   AddressMH[3].Ref_PLC_set_value_CP := 0;
   AddressMH[3].Ref_NozzelBypassControl := 0;
   AddressMH[3].Ref_NozzelBypassSetOut := 0;
   AddressMH[3].Ref_Reserve := 0;
   AddressMH[3].Ref_OK := FALSE;
   AddressMH[3].MH_Channel_01 := TRUE;
   AddressMH[3].MH_Channel_02 := FALSE;
   AddressMH[3].Spare_03 := FALSE;
   AddressMH[3].Spare_04 := FALSE;
   AddressMH[3].Spare_05 := FALSE;
   AddressMH[3].Spare_06 := FALSE;
   AddressMH[3].Spare_07 := FALSE;
   AddressMH[4].Ref_Digital_Input := 32;
   AddressMH[4].Ref_MH_ShotTime := 1550;
   AddressMH[4].Ref_MH_Opening_Time := 1554;
   AddressMH[4].Ref_MH_Closing_Time := 1556;
   AddressMH[4].Ref_MH_State := 1560;
   AddressMH[4].Ref_PLC_State := 0;
   AddressMH[4].Ref_CP_State := 0;
   AddressMH[4].Ref_Digital_Output := 32;
   AddressMH[4].Ref_ShotTimeSetValue := 1550;
   AddressMH[4].Ref_ServiceProduction := 1554;
   AddressMH[4].Ref_MixingheadControl := 1560;
   AddressMH[4].Ref_PLC_comand_SP := 0;
   AddressMH[4].Ref_PLC_comand_CP := 0;
   AddressMH[4].Ref_PLC_set_value_SP := 0;
   AddressMH[4].Ref_PLC_set_value_CP := 0;
   AddressMH[4].Ref_NozzelBypassControl := 0;
   AddressMH[4].Ref_NozzelBypassSetOut := 0;
   AddressMH[4].Ref_Reserve := 0;
   AddressMH[4].Ref_OK := FALSE;
   AddressMH[4].MH_Channel_01 := TRUE;
   AddressMH[4].MH_Channel_02 := FALSE;
   AddressMH[4].Spare_03 := FALSE;
   AddressMH[4].Spare_04 := FALSE;
   AddressMH[4].Spare_05 := FALSE;
   AddressMH[4].Spare_06 := FALSE;
   AddressMH[4].Spare_07 := FALSE;
   AddressMH[5].Ref_Digital_Input := 36;
   AddressMH[5].Ref_MH_ShotTime := 1636;
   AddressMH[5].Ref_MH_Opening_Time := 1640;
   AddressMH[5].Ref_MH_Closing_Time := 1642;
   AddressMH[5].Ref_MH_State := 1644;
   AddressMH[5].Ref_PLC_State := 0;
   AddressMH[5].Ref_CP_State := 0;
   AddressMH[5].Ref_Digital_Output := 36;
   AddressMH[5].Ref_ShotTimeSetValue := 1636;
   AddressMH[5].Ref_ServiceProduction := 1640;
   AddressMH[5].Ref_MixingheadControl := 1642;
   AddressMH[5].Ref_PLC_comand_SP := 0;
   AddressMH[5].Ref_PLC_comand_CP := 0;
   AddressMH[5].Ref_PLC_set_value_SP := 0;
   AddressMH[5].Ref_PLC_set_value_CP := 0;
   AddressMH[5].Ref_NozzelBypassControl := 0;
   AddressMH[5].Ref_NozzelBypassSetOut := 0;
   AddressMH[5].Ref_Reserve := 0;
   AddressMH[5].Ref_OK := FALSE;
   AddressMH[5].MH_Channel_01 := TRUE;
   AddressMH[5].MH_Channel_02 := FALSE;
   AddressMH[5].Spare_03 := FALSE;
   AddressMH[5].Spare_04 := FALSE;
   AddressMH[5].Spare_05 := FALSE;
   AddressMH[5].Spare_06 := FALSE;
   AddressMH[5].Spare_07 := FALSE;
   AddressMH[6].Ref_Digital_Input := 40;
   AddressMH[6].Ref_MH_ShotTime := 1686;
   AddressMH[6].Ref_MH_Opening_Time := 1690;
   AddressMH[6].Ref_MH_Closing_Time := 1692;
   AddressMH[6].Ref_MH_State := 1694;
   AddressMH[6].Ref_PLC_State := 0;
   AddressMH[6].Ref_CP_State := 0;
   AddressMH[6].Ref_Digital_Output := 40;
   AddressMH[6].Ref_ShotTimeSetValue := 1686;
   AddressMH[6].Ref_ServiceProduction := 1690;
   AddressMH[6].Ref_MixingheadControl := 1692;
   AddressMH[6].Ref_PLC_comand_SP := 0;
   AddressMH[6].Ref_PLC_comand_CP := 0;
   AddressMH[6].Ref_PLC_set_value_SP := 0;
   AddressMH[6].Ref_PLC_set_value_CP := 0;
   AddressMH[6].Ref_NozzelBypassControl := 0;
   AddressMH[6].Ref_NozzelBypassSetOut := 0;
   AddressMH[6].Ref_Reserve := 0;
   AddressMH[6].Ref_OK := FALSE;
   AddressMH[6].MH_Channel_01 := TRUE;
   AddressMH[6].MH_Channel_02 := FALSE;
   AddressMH[6].Spare_03 := FALSE;
   AddressMH[6].Spare_04 := FALSE;
   AddressMH[6].Spare_05 := FALSE;
   AddressMH[6].Spare_06 := FALSE;
   AddressMH[6].Spare_07 := FALSE;
   AddressMH[7].Ref_Digital_Input := 44;
   AddressMH[7].Ref_MH_ShotTime := 1736;
   AddressMH[7].Ref_MH_Opening_Time := 1740;
   AddressMH[7].Ref_MH_Closing_Time := 1742;
   AddressMH[7].Ref_MH_State := 1744;
   AddressMH[7].Ref_PLC_State := 0;
   AddressMH[7].Ref_CP_State := 0;
   AddressMH[7].Ref_Digital_Output := 44;
   AddressMH[7].Ref_ShotTimeSetValue := 1736;
   AddressMH[7].Ref_ServiceProduction := 1740;
   AddressMH[7].Ref_MixingheadControl := 1742;
   AddressMH[7].Ref_PLC_comand_SP := 0;
   AddressMH[7].Ref_PLC_comand_CP := 0;
   AddressMH[7].Ref_PLC_set_value_SP := 0;
   AddressMH[7].Ref_PLC_set_value_CP := 0;
   AddressMH[7].Ref_NozzelBypassControl := 0;
   AddressMH[7].Ref_NozzelBypassSetOut := 0;
   AddressMH[7].Ref_Reserve := 0;
   // 242 more start values not shown
END_DATA_BLOCK

DATA_BLOCK "DB1233_ProCanIO_Flow"   // DB1233
TITLE = Address allocation flow IO-ProCan
{ S7_Optimized_Access := 'FALSE' }
VERSION : 0.1
   VAR
      ReadWriteDeviceNo : Int := 1;
      CopyDeviceNO : Int := 0;
      Read : Bool := FALSE;
      Write : Bool := FALSE;
      Copy : Bool := FALSE;
      AddressFlow : Array[0..16] of "UDT1233_ProCanIO_Flow";
   END_VAR
BEGIN
   AddressFlow[1].Ref_Act_FlowValue := 2000;
   AddressFlow[2].Ref_Act_FlowValue := 2004;
   AddressFlow[3].Ref_Act_FlowValue := 800;
   AddressFlow[4].Ref_Act_FlowValue := 0;
   AddressFlow[5].Ref_Act_FlowValue := 0;
   AddressFlow[6].Ref_Act_FlowValue := 0;
   AddressFlow[7].Ref_Act_FlowValue := 0;
   AddressFlow[8].Ref_Act_FlowValue := 0;
   AddressFlow[9].Ref_Act_FlowValue := 0;
   AddressFlow[10].Ref_Act_FlowValue := 0;
   AddressFlow[11].Ref_Act_FlowValue := 0;
   AddressFlow[12].Ref_Act_FlowValue := 0;
   AddressFlow[1].Ref_Act_FlowState := 2032;
   AddressFlow[2].Ref_Act_FlowState := 2033;
   AddressFlow[3].Ref_Act_FlowState := 0;
   AddressFlow[4].Ref_Act_FlowState := 0;
   AddressFlow[5].Ref_Act_FlowState := 0;
   AddressFlow[6].Ref_Act_FlowState := 0;
   AddressFlow[7].Ref_Act_FlowState := 0;
   AddressFlow[8].Ref_Act_FlowState := 0;
   AddressFlow[9].Ref_Act_FlowState := 0;
   AddressFlow[10].Ref_Act_FlowState := 0;
   AddressFlow[11].Ref_Act_FlowState := 0;
   AddressFlow[12].Ref_Act_FlowState := 0;
   AddressFlow[1].Ref_Set_FlowRate := 2000;
   AddressFlow[2].Ref_Set_FlowRate := 2004;
   AddressFlow[3].Ref_Set_FlowRate := 0;
   AddressFlow[4].Ref_Set_FlowRate := 0;
   AddressFlow[5].Ref_Set_FlowRate := 0;
   AddressFlow[6].Ref_Set_FlowRate := 0;
   AddressFlow[7].Ref_Set_FlowRate := 0;
   AddressFlow[8].Ref_Set_FlowRate := 0;
   AddressFlow[9].Ref_Set_FlowRate := 0;
   AddressFlow[10].Ref_Set_FlowRate := 0;
   AddressFlow[11].Ref_Set_FlowRate := 0;
   AddressFlow[12].Ref_Set_FlowRate := 0;
   AddressFlow[1].Ref_Set_FlowRateQPB := 2016;
   AddressFlow[2].Ref_Set_FlowRateQPB := 2020;
   AddressFlow[3].Ref_Set_FlowRateQPB := 0;
   AddressFlow[4].Ref_Set_FlowRateQPB := 0;
   AddressFlow[5].Ref_Set_FlowRateQPB := 0;
   AddressFlow[6].Ref_Set_FlowRateQPB := 0;
   AddressFlow[7].Ref_Set_FlowRateQPB := 0;
   AddressFlow[8].Ref_Set_FlowRateQPB := 0;
   AddressFlow[9].Ref_Set_FlowRateQPB := 0;
   AddressFlow[10].Ref_Set_FlowRateQPB := 0;
   AddressFlow[11].Ref_Set_FlowRateQPB := 0;
   AddressFlow[12].Ref_Set_FlowRateQPB := 0;
   AddressFlow[1].Ref_Set_SWO_PressureQPB := 2032;
   AddressFlow[2].Ref_Set_SWO_PressureQPB := 2034;
   AddressFlow[3].Ref_Set_SWO_PressureQPB := 0;
   AddressFlow[4].Ref_Set_SWO_PressureQPB := 0;
   AddressFlow[5].Ref_Set_SWO_PressureQPB := 0;
   AddressFlow[6].Ref_Set_SWO_PressureQPB := 0;
   AddressFlow[7].Ref_Set_SWO_PressureQPB := 0;
   AddressFlow[8].Ref_Set_SWO_PressureQPB := 0;
   AddressFlow[9].Ref_Set_SWO_PressureQPB := 0;
   AddressFlow[10].Ref_Set_SWO_PressureQPB := 0;
   AddressFlow[11].Ref_Set_SWO_PressureQPB := 0;
   AddressFlow[12].Ref_Set_SWO_PressureQPB := 0;
   AddressFlow[1].Ref_Set_FlowIndexFlags := 2040;
   AddressFlow[2].Ref_Set_FlowIndexFlags := 2041;
   AddressFlow[3].Ref_Set_FlowIndexFlags := 0;
   AddressFlow[4].Ref_Set_FlowIndexFlags := 0;
   AddressFlow[5].Ref_Set_FlowIndexFlags := 0;
   AddressFlow[6].Ref_Set_FlowIndexFlags := 0;
   AddressFlow[7].Ref_Set_FlowIndexFlags := 0;
   AddressFlow[8].Ref_Set_FlowIndexFlags := 0;
   AddressFlow[9].Ref_Set_FlowIndexFlags := 0;
   AddressFlow[10].Ref_Set_FlowIndexFlags := 0;
   AddressFlow[11].Ref_Set_FlowIndexFlags := 0;
   AddressFlow[12].Ref_Set_FlowIndexFlags := 0;
   AddressFlow[1].Ref_PistonPosition := 0;
   AddressFlow[7].Ref_PistonPosition := 0;
   AddressFlow[1].Ref_OK := TRUE;
   AddressFlow[2].Ref_OK := TRUE;
   AddressFlow[3].Ref_OK := FALSE;
   AddressFlow[4].Ref_OK := FALSE;
   AddressFlow[5].Ref_OK := FALSE;
   AddressFlow[6].Ref_OK := FALSE;
   AddressFlow[7].Ref_OK := FALSE;
   AddressFlow[8].Ref_OK := FALSE;
   AddressFlow[9].Ref_OK := FALSE;
   AddressFlow[10].Ref_OK := FALSE;
   AddressFlow[11].Ref_OK := FALSE;
   AddressFlow[12].Ref_OK := FALSE;
   AddressFlow[3].Ref_Act_PressureQPB := 0;
   AddressFlow[3].Ref_TandemStatus := 0;
   AddressFlow[0].Ref_Act_FlowValue := 2000;
   AddressFlow[0].Ref_Act_FlowState := 2032;
   AddressFlow[0].Ref_Set_FlowRate := 2000;
   AddressFlow[0].Ref_Set_FlowRateQPB := 2016;
   AddressFlow[0].Ref_Act_PressureQPB := 0;
   AddressFlow[0].Ref_Set_SWO_PressureQPB := 2032;
   AddressFlow[0].Ref_Set_FlowIndexFlags := 2040;
   AddressFlow[0].Ref_TandemStatus := 0;
   AddressFlow[0].Ref_TandemComand := 0;
   AddressFlow[0].Ref_PistonPosition := 0;
   AddressFlow[0].Ref_OK := TRUE;
   AddressFlow[1].Ref_Act_PressureQPB := 0;
   AddressFlow[1].Ref_TandemStatus := 0;
   AddressFlow[1].Ref_TandemComand := 0;
   AddressFlow[2].Ref_Act_PressureQPB := 0;
   AddressFlow[2].Ref_TandemStatus := 0;
   AddressFlow[2].Ref_TandemComand := 0;
   AddressFlow[2].Ref_PistonPosition := 0;
   AddressFlow[3].Ref_TandemComand := 0;
   AddressFlow[3].Ref_PistonPosition := 0;
   AddressFlow[4].Ref_Act_PressureQPB := 0;
   AddressFlow[4].Ref_TandemStatus := 0;
   AddressFlow[4].Ref_TandemComand := 0;
   AddressFlow[4].Ref_PistonPosition := 0;
   AddressFlow[5].Ref_Act_PressureQPB := 0;
   AddressFlow[5].Ref_TandemStatus := 0;
   AddressFlow[5].Ref_TandemComand := 0;
   AddressFlow[5].Ref_PistonPosition := 0;
   AddressFlow[6].Ref_Act_PressureQPB := 0;
   AddressFlow[6].Ref_TandemStatus := 0;
   AddressFlow[6].Ref_TandemComand := 0;
   AddressFlow[6].Ref_PistonPosition := 0;
   AddressFlow[7].Ref_Act_PressureQPB := 0;
   AddressFlow[7].Ref_TandemStatus := 0;
   AddressFlow[7].Ref_TandemComand := 0;
   AddressFlow[8].Ref_Act_PressureQPB := 0;
   AddressFlow[8].Ref_TandemStatus := 0;
   AddressFlow[8].Ref_TandemComand := 0;
   AddressFlow[8].Ref_PistonPosition := 0;
   AddressFlow[9].Ref_Act_PressureQPB := 0;
   AddressFlow[9].Ref_TandemStatus := 0;
   AddressFlow[9].Ref_TandemComand := 0;
   AddressFlow[9].Ref_PistonPosition := 0;
   AddressFlow[10].Ref_Act_PressureQPB := 0;
   AddressFlow[10].Ref_TandemStatus := 0;
   AddressFlow[10].Ref_TandemComand := 0;
   AddressFlow[10].Ref_PistonPosition := 0;
   AddressFlow[11].Ref_Act_PressureQPB := 0;
   AddressFlow[11].Ref_TandemStatus := 0;
   AddressFlow[11].Ref_TandemComand := 0;
   AddressFlow[11].Ref_PistonPosition := 0;
   AddressFlow[12].Ref_Act_PressureQPB := 0;
   AddressFlow[12].Ref_TandemStatus := 0;
   AddressFlow[12].Ref_TandemComand := 0;
   AddressFlow[12].Ref_PistonPosition := 0;
   AddressFlow[13].Ref_Act_FlowValue := 0;
   AddressFlow[13].Ref_Act_FlowState := 0;
   AddressFlow[13].Ref_Set_FlowRate := 0;
   AddressFlow[13].Ref_Set_FlowRateQPB := 0;
   AddressFlow[13].Ref_Act_PressureQPB := 0;
   AddressFlow[13].Ref_Set_SWO_PressureQPB := 0;
   AddressFlow[13].Ref_Set_FlowIndexFlags := 0;
   AddressFlow[13].Ref_TandemStatus := 0;
   AddressFlow[13].Ref_TandemComand := 0;
   AddressFlow[13].Ref_PistonPosition := 0;
   AddressFlow[13].Ref_OK := FALSE;
   AddressFlow[14].Ref_Act_FlowValue := 0;
   AddressFlow[14].Ref_Act_FlowState := 0;
   AddressFlow[14].Ref_Set_FlowRate := 0;
   AddressFlow[14].Ref_Set_FlowRateQPB := 0;
   AddressFlow[14].Ref_Act_PressureQPB := 0;
   AddressFlow[14].Ref_Set_SWO_PressureQPB := 0;
   AddressFlow[14].Ref_Set_FlowIndexFlags := 0;
   AddressFlow[14].Ref_TandemStatus := 0;
   AddressFlow[14].Ref_TandemComand := 0;
   AddressFlow[14].Ref_PistonPosition := 0;
   AddressFlow[14].Ref_OK := FALSE;
   AddressFlow[15].Ref_Act_FlowValue := 0;
   AddressFlow[15].Ref_Act_FlowState := 0;
   AddressFlow[15].Ref_Set_FlowRate := 0;
   AddressFlow[15].Ref_Set_FlowRateQPB := 0;
   AddressFlow[15].Ref_Act_PressureQPB := 0;
   AddressFlow[15].Ref_Set_SWO_PressureQPB := 0;
   AddressFlow[15].Ref_Set_FlowIndexFlags := 0;
   AddressFlow[15].Ref_TandemStatus := 0;
   AddressFlow[15].Ref_TandemComand := 0;
   AddressFlow[15].Ref_PistonPosition := 0;
   AddressFlow[15].Ref_OK := FALSE;
   AddressFlow[16].Ref_Act_FlowValue := 0;
   AddressFlow[16].Ref_Act_FlowState := 0;
   AddressFlow[16].Ref_Set_FlowRate := 0;
   AddressFlow[16].Ref_Set_FlowRateQPB := 0;
   AddressFlow[16].Ref_Act_PressureQPB := 0;
   AddressFlow[16].Ref_Set_SWO_PressureQPB := 0;
   AddressFlow[16].Ref_Set_FlowIndexFlags := 0;
   AddressFlow[16].Ref_TandemStatus := 0;
   AddressFlow[16].Ref_TandemComand := 0;
   AddressFlow[16].Ref_PistonPosition := 0;
   AddressFlow[16].Ref_OK := FALSE;
END_DATA_BLOCK

DATA_BLOCK "DB1500_ShotDataToMC"   // DB1500
{ S7_Optimized_Access := 'FALSE' }
VERSION : 0.1
   VAR
      ShotData_MC : Array[0..4] of "ShotDataToMC";
   END_VAR
BEGIN
END_DATA_BLOCK

DATA_BLOCK "DB1900_IF_Robots"   // DB1900
{ S7_Optimized_Access := 'FALSE' }
VERSION : 0.1
   VAR
      ReadWriteDeviceNo : Int := 1;
      CopyDeviceNO : Int := 0;
      Read : Bool := FALSE;
      Write : Bool := FALSE;
      Copy : Bool := FALSE;
      Switch_Robots : Array[0..4] of Struct   // Switch Robots / State Robots
         SwitchHomePosON_OFF : Bool;
         SwitchMaintPosON_OFF : Bool;
         SwitchMaintPos_2ON_OFF : Bool;
         SwitchTestShotON_OFF : Bool;
         SwitchCleaningON_OFF : Bool;
         SwitchBrushON_OFF : Bool;
         SwitchSyncON_OFF : Bool;
         SwitchTeachenON_OFF : Bool;
         SwitchLearningON_OFF : Bool;
         SwitchAirCleaningON_OFF : Bool;
         SwitchAirCleaningManON_OFF : Bool;
         SwitchSpare_12 : Bool;
         SwitchSpare_13 : Bool;
         SwitchSpare_14 : Bool;
         SwitchSpare_15 : Bool;
         SwitchSpare_16 : Bool;
         StateHomePos : Byte;
         StateMaintPos : Byte;
         StateMaintPos_2 : Byte;
         StateTestShot : Byte;
         StateCleaning : Byte;
         StateBrush : Byte;
         StateSync : Byte;
         StateTeachen : Byte;
         StateLearning : Byte;
         StateAirCleaning : Byte;
         StateAirCleaningManual : Byte;
         State_12 : Byte;
         State_13 : Byte;
         State_14 : Byte;
         State_15 : Byte;
         State_16 : Byte;
      END_STRUCT;
      State_Robots : Array[0..4] of Struct   // State Robots for HMI
         Rob_in_Home : Bool;
         Rob_in_Automatic : Bool;
         Rob_in_Cycle : Bool;
         Fault_Exist : Bool;
         EmergencyStopReady : Bool;
         AutomatcStopReady : Bool;
         MixingheadAuto : Bool;
         MaschineAuto : Bool;
         CleaningMHRequested : Bool;
         CleaningMHOn : Bool;
         ReadyForStartCycle : Bool;
         TestShotRunning : Bool;
         AtPos1or2 : Bool;   // Die Schnittstellen an diesen Roboter sind an erster oder zweiter Stelle angemeldet
         Spare_1_5 : Bool;
         Spare_1_6 : Bool;
         Spare_1_7 : Bool;
         Rob_Prog_No : Byte;
         Rob_MC_No : Byte;
         StepNo : Byte;
         FaultNo : Byte;
         Spare_6 : Byte;
         Spare_7 : Byte;
         Spare_8 : Byte;
      END_STRUCT;
      Faults_Robots : Array[0..4] of "General_Faults";   // Faults Robots for HMI
      State_Kuka : Array[0..4] of "Kuka_KRC4_Status";   // State/Input/Ouput Kuka
      State_ABB : Array[0..4] of "ABB_IRC6_State";   // State/Input/Ouput ABB
      State_Fanuc : Array[0..4] of "Fanuc_Status";   // State/Input/Ouput Fanuc
   END_VAR
BEGIN
   Switch_Robots[0].SwitchHomePosON_OFF := FALSE;
   Switch_Robots[0].SwitchMaintPosON_OFF := FALSE;
   Switch_Robots[0].SwitchMaintPos_2ON_OFF := FALSE;
   Switch_Robots[0].SwitchTestShotON_OFF := FALSE;
   Switch_Robots[0].SwitchCleaningON_OFF := FALSE;
   Switch_Robots[0].SwitchBrushON_OFF := FALSE;
   Switch_Robots[0].SwitchSyncON_OFF := FALSE;
   Switch_Robots[0].SwitchTeachenON_OFF := FALSE;
   Switch_Robots[0].SwitchLearningON_OFF := FALSE;
   Switch_Robots[0].SwitchAirCleaningON_OFF := FALSE;
   Switch_Robots[0].SwitchAirCleaningManON_OFF := FALSE;
   Switch_Robots[0].SwitchSpare_12 := FALSE;
   Switch_Robots[0].SwitchSpare_13 := FALSE;
   Switch_Robots[0].SwitchSpare_14 := FALSE;
   Switch_Robots[0].SwitchSpare_15 := FALSE;
   Switch_Robots[0].SwitchSpare_16 := FALSE;
   Switch_Robots[0].StateHomePos := 16#00;
   Switch_Robots[0].StateMaintPos := 16#00;
   Switch_Robots[0].StateMaintPos_2 := 16#00;
   Switch_Robots[0].StateTestShot := 16#00;
   Switch_Robots[0].StateCleaning := 16#00;
   Switch_Robots[0].StateBrush := 16#00;
   Switch_Robots[0].StateSync := 16#02;
   Switch_Robots[0].StateTeachen := 16#00;
   Switch_Robots[0].StateLearning := 16#00;
   Switch_Robots[0].StateAirCleaning := 16#00;
   Switch_Robots[0].StateAirCleaningManual := 16#00;
   Switch_Robots[0].State_12 := 16#00;
   Switch_Robots[0].State_13 := 16#00;
   Switch_Robots[0].State_14 := 16#00;
   Switch_Robots[0].State_15 := 16#00;
   Switch_Robots[0].State_16 := 16#00;
   Switch_Robots[1].SwitchHomePosON_OFF := FALSE;
   Switch_Robots[1].SwitchMaintPosON_OFF := FALSE;
   Switch_Robots[1].SwitchMaintPos_2ON_OFF := FALSE;
   Switch_Robots[1].SwitchTestShotON_OFF := FALSE;
   Switch_Robots[1].SwitchCleaningON_OFF := FALSE;
   Switch_Robots[1].SwitchBrushON_OFF := FALSE;
   Switch_Robots[1].SwitchSyncON_OFF := FALSE;
   Switch_Robots[1].SwitchTeachenON_OFF := FALSE;
   Switch_Robots[1].SwitchLearningON_OFF := FALSE;
   Switch_Robots[1].SwitchAirCleaningON_OFF := FALSE;
   Switch_Robots[1].SwitchAirCleaningManON_OFF := FALSE;
   Switch_Robots[1].SwitchSpare_12 := FALSE;
   Switch_Robots[1].SwitchSpare_13 := FALSE;
   Switch_Robots[1].SwitchSpare_14 := FALSE;
   Switch_Robots[1].SwitchSpare_15 := FALSE;
   Switch_Robots[1].SwitchSpare_16 := FALSE;
   Switch_Robots[1].StateHomePos := 16#00;
   Switch_Robots[1].StateMaintPos := 16#00;
   Switch_Robots[1].StateMaintPos_2 := 16#00;
   Switch_Robots[1].StateTestShot := 16#00;
   Switch_Robots[1].StateCleaning := 16#00;
   Switch_Robots[1].StateBrush := 16#00;
   Switch_Robots[1].StateSync := 16#02;
   Switch_Robots[1].StateTeachen := 16#00;
   Switch_Robots[1].StateLearning := 16#00;
   Switch_Robots[1].StateAirCleaning := 16#00;
   Switch_Robots[1].StateAirCleaningManual := 16#00;
   Switch_Robots[1].State_12 := 16#00;
   Switch_Robots[1].State_13 := 16#00;
   Switch_Robots[1].State_14 := 16#00;
   Switch_Robots[1].State_15 := 16#00;
   Switch_Robots[1].State_16 := 16#00;
   Switch_Robots[2].SwitchHomePosON_OFF := FALSE;
   Switch_Robots[2].SwitchMaintPosON_OFF := FALSE;
   Switch_Robots[2].SwitchMaintPos_2ON_OFF := FALSE;
   Switch_Robots[2].SwitchTestShotON_OFF := FALSE;
   Switch_Robots[2].SwitchCleaningON_OFF := FALSE;
   Switch_Robots[2].SwitchBrushON_OFF := FALSE;
   Switch_Robots[2].SwitchSyncON_OFF := FALSE;
   Switch_Robots[2].SwitchTeachenON_OFF := FALSE;
   Switch_Robots[2].SwitchLearningON_OFF := FALSE;
   Switch_Robots[2].SwitchAirCleaningON_OFF := FALSE;
   Switch_Robots[2].SwitchAirCleaningManON_OFF := FALSE;
   Switch_Robots[2].SwitchSpare_12 := FALSE;
   Switch_Robots[2].SwitchSpare_13 := FALSE;
   Switch_Robots[2].SwitchSpare_14 := FALSE;
   Switch_Robots[2].SwitchSpare_15 := FALSE;
   Switch_Robots[2].SwitchSpare_16 := FALSE;
   Switch_Robots[2].StateHomePos := 16#00;
   Switch_Robots[2].StateMaintPos := 16#00;
   Switch_Robots[2].StateMaintPos_2 := 16#00;
   Switch_Robots[2].StateTestShot := 16#00;
   Switch_Robots[2].StateCleaning := 16#00;
   Switch_Robots[2].StateBrush := 16#00;
   Switch_Robots[2].StateSync := 16#00;
   Switch_Robots[2].StateTeachen := 16#00;
   Switch_Robots[2].StateLearning := 16#00;
   Switch_Robots[2].StateAirCleaning := 16#00;
   Switch_Robots[2].StateAirCleaningManual := 16#00;
   Switch_Robots[2].State_12 := 16#00;
   Switch_Robots[2].State_13 := 16#00;
   Switch_Robots[2].State_14 := 16#00;
   Switch_Robots[2].State_15 := 16#00;
   Switch_Robots[2].State_16 := 16#00;
   Switch_Robots[3].SwitchHomePosON_OFF := FALSE;
   Switch_Robots[3].SwitchMaintPosON_OFF := FALSE;
   Switch_Robots[3].SwitchMaintPos_2ON_OFF := FALSE;
   Switch_Robots[3].SwitchTestShotON_OFF := FALSE;
   Switch_Robots[3].SwitchCleaningON_OFF := FALSE;
   Switch_Robots[3].SwitchBrushON_OFF := FALSE;
   Switch_Robots[3].SwitchSyncON_OFF := FALSE;
   Switch_Robots[3].SwitchTeachenON_OFF := FALSE;
   Switch_Robots[3].SwitchLearningON_OFF := FALSE;
   Switch_Robots[3].SwitchAirCleaningON_OFF := FALSE;
   Switch_Robots[3].SwitchAirCleaningManON_OFF := FALSE;
   Switch_Robots[3].SwitchSpare_12 := FALSE;
   Switch_Robots[3].SwitchSpare_13 := FALSE;
   Switch_Robots[3].SwitchSpare_14 := FALSE;
   Switch_Robots[3].SwitchSpare_15 := FALSE;
   Switch_Robots[3].SwitchSpare_16 := FALSE;
   Switch_Robots[3].StateHomePos := 16#00;
   Switch_Robots[3].StateMaintPos := 16#00;
   Switch_Robots[3].StateMaintPos_2 := 16#00;
   Switch_Robots[3].StateTestShot := 16#00;
   Switch_Robots[3].StateCleaning := 16#00;
   Switch_Robots[3].StateBrush := 16#00;
   Switch_Robots[3].StateSync := 16#00;
   Switch_Robots[3].StateTeachen := 16#00;
   Switch_Robots[3].StateLearning := 16#00;
   Switch_Robots[3].StateAirCleaning := 16#00;
   Switch_Robots[3].StateAirCleaningManual := 16#00;
   Switch_Robots[3].State_12 := 16#00;
   Switch_Robots[3].State_13 := 16#00;
   Switch_Robots[3].State_14 := 16#00;
   Switch_Robots[3].State_15 := 16#00;
   Switch_Robots[3].State_16 := 16#00;
   Switch_Robots[4].SwitchHomePosON_OFF := FALSE;
   Switch_Robots[4].SwitchMaintPosON_OFF := FALSE;
   Switch_Robots[4].SwitchMaintPos_2ON_OFF := FALSE;
   Switch_Robots[4].SwitchTestShotON_OFF := FALSE;
   Switch_Robots[4].SwitchCleaningON_OFF := FALSE;
   Switch_Robots[4].SwitchBrushON_OFF := FALSE;
   Switch_Robots[4].SwitchSyncON_OFF := FALSE;
   Switch_Robots[4].SwitchTeachenON_OFF := FALSE;
   Switch_Robots[4].SwitchLearningON_OFF := FALSE;
   Switch_Robots[4].SwitchAirCleaningON_OFF := FALSE;
   Switch_Robots[4].SwitchAirCleaningManON_OFF := FALSE;
   Switch_Robots[4].SwitchSpare_12 := FALSE;
   Switch_Robots[4].SwitchSpare_13 := FALSE;
   Switch_Robots[4].SwitchSpare_14 := FALSE;
   Switch_Robots[4].SwitchSpare_15 := FALSE;
   Switch_Robots[4].SwitchSpare_16 := FALSE;
   Switch_Robots[4].StateHomePos := 16#00;
   Switch_Robots[4].StateMaintPos := 16#00;
   Switch_Robots[4].StateMaintPos_2 := 16#00;
   Switch_Robots[4].StateTestShot := 16#00;
   Switch_Robots[4].StateCleaning := 16#00;
   Switch_Robots[4].StateBrush := 16#00;
   Switch_Robots[4].StateSync := 16#00;
   Switch_Robots[4].StateTeachen := 16#00;
   Switch_Robots[4].StateLearning := 16#00;
   Switch_Robots[4].StateAirCleaning := 16#00;
   Switch_Robots[4].StateAirCleaningManual := 16#00;
   Switch_Robots[4].State_12 := 16#00;
   Switch_Robots[4].State_13 := 16#00;
   Switch_Robots[4].State_14 := 16#00;
   Switch_Robots[4].State_15 := 16#00;
   Switch_Robots[4].State_16 := 16#00;
   State_Robots[0].Rob_in_Home := FALSE;
   State_Robots[0].Rob_in_Automatic := FALSE;
   State_Robots[0].Rob_in_Cycle := FALSE;
   State_Robots[0].Fault_Exist := FALSE;
   State_Robots[0].EmergencyStopReady := TRUE;
   State_Robots[0].AutomatcStopReady := TRUE;
   State_Robots[0].MixingheadAuto := FALSE;
   State_Robots[0].MaschineAuto := FALSE;
   State_Robots[0].CleaningMHRequested := TRUE;
   State_Robots[0].CleaningMHOn := FALSE;
   State_Robots[0].ReadyForStartCycle := FALSE;
   State_Robots[0].TestShotRunning := FALSE;
   State_Robots[0].AtPos1or2 := FALSE;
   State_Robots[0].Spare_1_5 := FALSE;
   State_Robots[0].Spare_1_6 := FALSE;
   State_Robots[0].Spare_1_7 := FALSE;
   State_Robots[0].Rob_Prog_No := 16#00;
   State_Robots[0].Rob_MC_No := 16#00;
   State_Robots[0].StepNo := 16#00;
   State_Robots[0].FaultNo := 16#00;
   State_Robots[0].Spare_6 := 16#00;
   State_Robots[0].Spare_7 := 16#00;
   State_Robots[0].Spare_8 := 16#00;
   State_Robots[1].Rob_in_Home := FALSE;
   State_Robots[1].Rob_in_Automatic := FALSE;
   State_Robots[1].Rob_in_Cycle := FALSE;
   State_Robots[1].Fault_Exist := FALSE;
   State_Robots[1].EmergencyStopReady := FALSE;
   State_Robots[1].AutomatcStopReady := FALSE;
   State_Robots[1].MixingheadAuto := FALSE;
   State_Robots[1].MaschineAuto := FALSE;
   State_Robots[1].CleaningMHRequested := TRUE;
   State_Robots[1].CleaningMHOn := FALSE;
   State_Robots[1].ReadyForStartCycle := FALSE;
   State_Robots[1].TestShotRunning := FALSE;
   State_Robots[1].AtPos1or2 := FALSE;
   State_Robots[1].Spare_1_5 := FALSE;
   State_Robots[1].Spare_1_6 := FALSE;
   State_Robots[1].Spare_1_7 := FALSE;
   State_Robots[1].Rob_Prog_No := 16#00;
   // 3950 more start values not shown
END_DATA_BLOCK

